   4910: 'Spare_Fault_4910', class No Acknowledgement, trigger "DB302_HMI_Faults_Carrier76_Faults_2" bit 13
   4911: 'Spare_Fault_4911', class No Acknowledgement, trigger "DB302_HMI_Faults_Carrier76_Faults_2" bit 14
   4912: 'Spare_Fault_4912', class No Acknowledgement, trigger "DB302_HMI_Faults_Carrier76_Faults_2" bit 15
   4913: 'Spare_Fault_4913', class No Acknowledgement, trigger "DB302_HMI_Faults_Carrier76_Faults_3" bit 0
   4914: 'Spare_Fault_4914', class No Acknowledgement, trigger "DB302_HMI_Faults_Carrier76_Faults_3" bit 1
   4915: 'Spare_Fault_4915', class No Acknowledgement, trigger "DB302_HMI_Faults_Carrier76_Faults_3" bit 2
   4916: 'Spare_Fault_4916', class No Acknowledgement, trigger "DB302_HMI_Faults_Carrier76_Faults_3" bit 3
   4917: 'Spare_Fault_4917', class No Acknowledgement, trigger "DB302_HMI_Faults_Carrier76_Faults_3" bit 4
   4918: 'Spare_Fault_4918', class No Acknowledgement, trigger "DB302_HMI_Faults_Carrier76_Faults_3" bit 5
   4919: 'Spare_Fault_4919', class No Acknowledgement, trigger "DB302_HMI_Faults_Carrier76_Faults_3" bit 6
   4920: 'Spare_Fault_4920', class No Acknowledgement, trigger "DB302_HMI_Faults_Carrier76_Faults_3" bit 7
   4921: 'Spare_Fault_4921', class No Acknowledgement, trigger "DB302_HMI_Faults_Carrier76_Faults_3" bit 8
   4922: 'Spare_Fault_4922', class No Acknowledgement, trigger "DB302_HMI_Faults_Carrier76_Faults_3" bit 9
   4923: 'Spare_Fault_4923', class No Acknowledgement, trigger "DB302_HMI_Faults_Carrier76_Faults_3" bit 10
   4924: 'Spare_Fault_4924', class No Acknowledgement, trigger "DB302_HMI_Faults_Carrier76_Faults_3" bit 11
   4925: 'Spare_Fault_4925', class No Acknowledgement, trigger "DB302_HMI_Faults_Carrier76_Faults_3" bit 12
   4926: 'Spare_Fault_4926', class No Acknowledgement, trigger "DB302_HMI_Faults_Carrier76_Faults_3" bit 13
   4927: 'Spare_Fault_4927', class No Acknowledgement, trigger "DB302_HMI_Faults_Carrier76_Faults_3" bit 14
   4928: 'Spare_Fault_4928', class No Acknowledgement, trigger "DB302_HMI_Faults_Carrier76_Faults_3" bit 15
   4929: 'Carrier 77 Disconnect Open Power Fault DI11.0', class No Acknowledgement, trigger "DB302_HMI_Faults_Carrier77_Faults_0" bit 0
   4930: 'Carrier 77 Drive Profinet Comm Fault', class No Acknowledgement, trigger "DB302_HMI_Faults_Carrier77_Faults_0" bit 1
   4931: 'Carrier 77 Production Stop Not Reset', class No Acknowledgement, trigger "DB302_HMI_Faults_Carrier77_Faults_0" bit 2
   4932: 'Carrier 77 CB02122 Tripped', class No Acknowledgement, trigger "DB302_HMI_Faults_Carrier77_Faults_0" bit 3
   4933: 'Carrier 77 CB02123 Tripped', class No Acknowledgement, trigger "DB302_HMI_Faults_Carrier77_Faults_0" bit 4
   4934: 'Carrier 77 AUX1 CB Tripped', class No Acknowledgement, trigger "DB302_HMI_Faults_Carrier77_Faults_0" bit 5
   4935: 'Carrier 77 AUX2 CB Tripped', class No Acknowledgement, trigger "DB302_HMI_Faults_Carrier77_Faults_0" bit 6
   4936: 'Carrier 77 PLC Not Communicating', class No Acknowledgement, trigger "DB302_HMI_Faults_Carrier77_Faults_0" bit 7
   4937: 'Carrier 77 Safe Input Card Fault', class No Acknowledgement, trigger "DB302_HMI_Faults_Carrier77_Faults_0" bit 8
   4938: 'Carrier 77 Safe Output Card Fault', class No Acknowledgement, trigger "DB302_HMI_Faults_Carrier77_Faults_0" bit 9
   4939: 'Carrier 77 Standard Input Card Fault', class No Acknowledgement, trigger "DB302_HMI_Faults_Carrier77_Faults_0" bit 10
   4940: 'Carrier 77 Standard Output Card Fault', class No Acknowledgement, trigger "DB302_HMI_Faults_Carrier77_Faults_0" bit 11
   4941: 'Carrier 77 Encoder Position Fault', class No Acknowledgement, trigger "DB302_HMI_Faults_Carrier77_Faults_0" bit 12
   4942: 'Carrier 77 Encoder Internal Error', class No Acknowledgement, trigger "DB302_HMI_Faults_Carrier77_Faults_0" bit 13
   4943: 'Carrier 77 Encoder Comm Fault', class No Acknowledgement, trigger "DB302_HMI_Faults_Carrier77_Faults_0" bit 14
   4944: 'Carrier 77 HMI Comm Fault', class No Acknowledgement, trigger "DB302_HMI_Faults_Carrier77_Faults_0" bit 15
   4945: 'Carrier 77 Crash Detection Fault', class No Acknowledgement, trigger "DB302_HMI_Faults_Carrier77_Faults_1" bit 0
   4946: 'Carrier 77 Carrier Number Invalid', class No Acknowledgement, trigger "DB302_HMI_Faults_Carrier77_Faults_1" bit 1
   4947: 'Carrier 77 Drive: PROFINET configuration error', class No Acknowledgement, trigger "DB302_HMI_Faults_Carrier77_Faults_1" bit 2
   4948: 'Carrier 77 Drive: Error internal communications', class No Acknowledgement, trigger "DB302_HMI_Faults_Carrier77_Faults_1" bit 3
   4949: 'Carrier 77 Drive: Motor overtemperature', class No Acknowledgement, trigger "DB302_HMI_Faults_Carrier77_Faults_1" bit 4
   4950: 'Carrier 77 Drive: Motor overcurrent', class No Acknowledgement, trigger "DB302_HMI_Faults_Carrier77_Faults_1" bit 5
   4951: 'Carrier 77 Drive: Infeed or power unit not ready', class No Acknowledgement, trigger "DB302_HMI_Faults_Carrier77_Faults_1" bit 6
   4952: 'Carrier 77 Drive: Short-circuit/ground fault detected', class No Acknowledgement, trigger "DB302_HMI_Faults_Carrier77_Faults_1" bit 7
   4953: 'Carrier 77 Drive: PROFINET Setpoint timeout', class No Acknowledgement, trigger "DB302_HMI_Faults_Carrier77_Faults_1" bit 8
   4954: 'Carrier 77 Power unit: Overcurrent', class No Acknowledgement, trigger "DB302_HMI_Faults_Carrier77_Faults_1" bit 9
   4955: 'Carrier 77 Power unit: DC link voltage overvoltage', class No Acknowledgement, trigger "DB302_HMI_Faults_Carrier77_Faults_1" bit 10
   4956: 'Carrier 77 Power unit: DC link voltage undervoltage', class No Acknowledgement, trigger "DB302_HMI_Faults_Carrier77_Faults_1" bit 11
   4957: 'Carrier 77 Power unit: Line phase failure in main circuit', class No Acknowledgement, trigger "DB302_HMI_Faults_Carrier77_Faults_1" bit 12
   4958: 'Carrier 77 Power unit: Phase failure motor cable', class No Acknowledgement, trigger "DB302_HMI_Faults_Carrier77_Faults_1" bit 13
   4959: 'Carrier 77 Power unit: Ground fault', class No Acknowledgement, trigger "DB302_HMI_Faults_Carrier77_Faults_1" bit 14
   4960: 'Spare_Fault_4960', class No Acknowledgement, trigger "DB302_HMI_Faults_Carrier77_Faults_1" bit 15
   4961: 'Carrier 77 Motion Off Fault', class No Acknowledgement, trigger "DB302_HMI_Faults_Carrier77_Faults_2" bit 0
   4962: 'Carrier 77 Motion On Fault', class No Acknowledgement, trigger "DB302_HMI_Faults_Carrier77_Faults_2" bit 1
   4963: 'Carrier 77 Spacing Fault', class No Acknowledgement, trigger "DB302_HMI_Faults_Carrier77_Faults_2" bit 2
   4964: 'Carrier 77 Duplicate Carrier Number Fault', class No Acknowledgement, trigger "DB302_HMI_Faults_Carrier77_Faults_2" bit 3
   4965: 'Spare_Fault_4965', class No Acknowledgement, trigger "DB302_HMI_Faults_Carrier77_Faults_2" bit 4
   4966: 'Spare_Fault_4966', class No Acknowledgement, trigger "DB302_HMI_Faults_Carrier77_Faults_2" bit 5
   4967: 'Spare_Fault_4967', class No Acknowledgement, trigger "DB302_HMI_Faults_Carrier77_Faults_2" bit 6
   4968: 'Spare_Fault_4968', class No Acknowledgement, trigger "DB302_HMI_Faults_Carrier77_Faults_2" bit 7
   4969: 'Spare_Fault_4969', class No Acknowledgement, trigger "DB302_HMI_Faults_Carrier77_Faults_2" bit 8
   4970: 'Spare_Fault_4970', class No Acknowledgement, trigger "DB302_HMI_Faults_Carrier77_Faults_2" bit 9
   4971: 'Spare_Fault_4971', class No Acknowledgement, trigger "DB302_HMI_Faults_Carrier77_Faults_2" bit 10
   4972: 'Spare_Fault_4972', class No Acknowledgement, trigger "DB302_HMI_Faults_Carrier77_Faults_2" bit 11
   4973: 'Spare_Fault_4973', class No Acknowledgement, trigger "DB302_HMI_Faults_Carrier77_Faults_2" bit 12
   4974: 'Spare_Fault_4974', class No Acknowledgement, trigger "DB302_HMI_Faults_Carrier77_Faults_2" bit 13
   4975: 'Spare_Fault_4975', class No Acknowledgement, trigger "DB302_HMI_Faults_Carrier77_Faults_2" bit 14
   4976: 'Spare_Fault_4976', class No Acknowledgement, trigger "DB302_HMI_Faults_Carrier77_Faults_2" bit 15
   4977: 'Spare_Fault_4977', class No Acknowledgement, trigger "DB302_HMI_Faults_Carrier77_Faults_3" bit 0
   4978: 'Spare_Fault_4978', class No Acknowledgement, trigger "DB302_HMI_Faults_Carrier77_Faults_3" bit 1
   4979: 'Spare_Fault_4979', class No Acknowledgement, trigger "DB302_HMI_Faults_Carrier77_Faults_3" bit 2
   4980: 'Spare_Fault_4980', class No Acknowledgement, trigger "DB302_HMI_Faults_Carrier77_Faults_3" bit 3
   4981: 'Spare_Fault_4981', class No Acknowledgement, trigger "DB302_HMI_Faults_Carrier77_Faults_3" bit 4
   4982: 'Spare_Fault_4982', class No Acknowledgement, trigger "DB302_HMI_Faults_Carrier77_Faults_3" bit 5
   4983: 'Spare_Fault_4983', class No Acknowledgement, trigger "DB302_HMI_Faults_Carrier77_Faults_3" bit 6
   4984: 'Spare_Fault_4984', class No Acknowledgement, trigger "DB302_HMI_Faults_Carrier77_Faults_3" bit 7
   4985: 'Spare_Fault_4985', class No Acknowledgement, trigger "DB302_HMI_Faults_Carrier77_Faults_3" bit 8
   4986: 'Spare_Fault_4986', class No Acknowledgement, trigger "DB302_HMI_Faults_Carrier77_Faults_3" bit 9
   4987: 'Spare_Fault_4987', class No Acknowledgement, trigger "DB302_HMI_Faults_Carrier77_Faults_3" bit 10
   4988: 'Spare_Fault_4988', class No Acknowledgement, trigger "DB302_HMI_Faults_Carrier77_Faults_3" bit 11
   4989: 'Spare_Fault_4989', class No Acknowledgement, trigger "DB302_HMI_Faults_Carrier77_Faults_3" bit 12
   4990: 'Spare_Fault_4990', class No Acknowledgement, trigger "DB302_HMI_Faults_Carrier77_Faults_3" bit 13
   4991: 'Spare_Fault_4991', class No Acknowledgement, trigger "DB302_HMI_Faults_Carrier77_Faults_3" bit 14
   4992: 'Spare_Fault_4992', class No Acknowledgement, trigger "DB302_HMI_Faults_Carrier77_Faults_3" bit 15
   4993: 'Carrier 78 Disconnect Open Power Fault DI11.0', class No Acknowledgement, trigger "DB302_HMI_Faults_Carrier78_Faults_0" bit 0
   4994: 'Carrier 78 Drive Profinet Comm Fault', class No Acknowledgement, trigger "DB302_HMI_Faults_Carrier78_Faults_0" bit 1
   4995: 'Carrier 78 Production Stop Not Reset', class No Acknowledgement, trigger "DB302_HMI_Faults_Carrier78_Faults_0" bit 2
   4996: 'Carrier 78 CB02122 Tripped', class No Acknowledgement, trigger "DB302_HMI_Faults_Carrier78_Faults_0" bit 3
   4997: 'Carrier 78 CB02123 Tripped', class No Acknowledgement, trigger "DB302_HMI_Faults_Carrier78_Faults_0" bit 4
   4998: 'Carrier 78 AUX1 CB Tripped', class No Acknowledgement, trigger "DB302_HMI_Faults_Carrier78_Faults_0" bit 5
   4999: 'Carrier 78 AUX2 CB Tripped', class No Acknowledgement, trigger "DB302_HMI_Faults_Carrier78_Faults_0" bit 6
   5000: 'Carrier 78 PLC Not Communicating', class No Acknowledgement, trigger "DB302_HMI_Faults_Carrier78_Faults_0" bit 7
   5001: 'Carrier 78 Safe Input Card Fault', class No Acknowledgement, trigger "DB302_HMI_Faults_Carrier78_Faults_0" bit 8
   5002: 'Carrier 78 Safe Output Card Fault', class No Acknowledgement, trigger "DB302_HMI_Faults_Carrier78_Faults_0" bit 9
   5003: 'Carrier 78 Standard Input Card Fault', class No Acknowledgement, trigger "DB302_HMI_Faults_Carrier78_Faults_0" bit 10
   5004: 'Carrier 78 Standard Output Card Fault', class No Acknowledgement, trigger "DB302_HMI_Faults_Carrier78_Faults_0" bit 11
   5005: 'Carrier 78 Encoder Position Fault', class No Acknowledgement, trigger "DB302_HMI_Faults_Carrier78_Faults_0" bit 12
   5006: 'Carrier 78 Encoder Internal Error', class No Acknowledgement, trigger "DB302_HMI_Faults_Carrier78_Faults_0" bit 13
   5007: 'Carrier 78 Encoder Comm Fault', class No Acknowledgement, trigger "DB302_HMI_Faults_Carrier78_Faults_0" bit 14
   5008: 'Carrier 78 HMI Comm Fault', class No Acknowledgement, trigger "DB302_HMI_Faults_Carrier78_Faults_0" bit 15
   5009: 'Carrier 78 Crash Detection Fault', class No Acknowledgement, trigger "DB302_HMI_Faults_Carrier78_Faults_1" bit 0
   5010: 'Carrier 78 Carrier Number Invalid', class No Acknowledgement, trigger "DB302_HMI_Faults_Carrier78_Faults_1" bit 1
   5011: 'Carrier 78 Drive: PROFINET configuration error', class No Acknowledgement, trigger "DB302_HMI_Faults_Carrier78_Faults_1" bit 2
   5012: 'Carrier 78 Drive: Error internal communications', class No Acknowledgement, trigger "DB302_HMI_Faults_Carrier78_Faults_1" bit 3
   5013: 'Carrier 78 Drive: Motor overtemperature', class No Acknowledgement, trigger "DB302_HMI_Faults_Carrier78_Faults_1" bit 4
   5014: 'Carrier 78 Drive: Motor overcurrent', class No Acknowledgement, trigger "DB302_HMI_Faults_Carrier78_Faults_1" bit 5
   5015: 'Carrier 78 Drive: Infeed or power unit not ready', class No Acknowledgement, trigger "DB302_HMI_Faults_Carrier78_Faults_1" bit 6
   5016: 'Carrier 78 Drive: Short-circuit/ground fault detected', class No Acknowledgement, trigger "DB302_HMI_Faults_Carrier78_Faults_1" bit 7
   5017: 'Carrier 78 Drive: PROFINET Setpoint timeout', class No Acknowledgement, trigger "DB302_HMI_Faults_Carrier78_Faults_1" bit 8
   5018: 'Carrier 78 Power unit: Overcurrent', class No Acknowledgement, trigger "DB302_HMI_Faults_Carrier78_Faults_1" bit 9
   5019: 'Carrier 78 Power unit: DC link voltage overvoltage', class No Acknowledgement, trigger "DB302_HMI_Faults_Carrier78_Faults_1" bit 10
   5020: 'Carrier 78 Power unit: DC link voltage undervoltage', class No Acknowledgement, trigger "DB302_HMI_Faults_Carrier78_Faults_1" bit 11
   5021: 'Carrier 78 Power unit: Line phase failure in main circuit', class No Acknowledgement, trigger "DB302_HMI_Faults_Carrier78_Faults_1" bit 12
   5022: 'Carrier 78 Power unit: Phase failure motor cable', class No Acknowledgement, trigger "DB302_HMI_Faults_Carrier78_Faults_1" bit 13
   5023: 'Carrier 78 Power unit: Ground fault', class No Acknowledgement, trigger "DB302_HMI_Faults_Carrier78_Faults_1" bit 14
   5024: 'Spare_Fault_5024', class No Acknowledgement, trigger "DB302_HMI_Faults_Carrier78_Faults_1" bit 15
   5025: 'Carrier 78 Motion Off Fault', class No Acknowledgement, trigger "DB302_HMI_Faults_Carrier78_Faults_2" bit 0
   5026: 'Carrier 78 Motion On Fault', class No Acknowledgement, trigger "DB302_HMI_Faults_Carrier78_Faults_2" bit 1
   5027: 'Carrier 78 Spacing Fault', class No Acknowledgement, trigger "DB302_HMI_Faults_Carrier78_Faults_2" bit 2
   5028: 'Carrier 78 Duplicate Carrier Number Fault', class No Acknowledgement, trigger "DB302_HMI_Faults_Carrier78_Faults_2" bit 3
   5029: 'Spare_Fault_5029', class No Acknowledgement, trigger "DB302_HMI_Faults_Carrier78_Faults_2" bit 4
   5030: 'Spare_Fault_5030', class No Acknowledgement, trigger "DB302_HMI_Faults_Carrier78_Faults_2" bit 5
   5031: 'Spare_Fault_5031', class No Acknowledgement, trigger "DB302_HMI_Faults_Carrier78_Faults_2" bit 6
   5032: 'Spare_Fault_5032', class No Acknowledgement, trigger "DB302_HMI_Faults_Carrier78_Faults_2" bit 7
   5033: 'Spare_Fault_5033', class No Acknowledgement, trigger "DB302_HMI_Faults_Carrier78_Faults_2" bit 8
   5034: 'Spare_Fault_5034', class No Acknowledgement, trigger "DB302_HMI_Faults_Carrier78_Faults_2" bit 9
   5035: 'Spare_Fault_5035', class No Acknowledgement, trigger "DB302_HMI_Faults_Carrier78_Faults_2" bit 10
   5036: 'Spare_Fault_5036', class No Acknowledgement, trigger "DB302_HMI_Faults_Carrier78_Faults_2" bit 11
   5037: 'Spare_Fault_5037', class No Acknowledgement, trigger "DB302_HMI_Faults_Carrier78_Faults_2" bit 12
   5038: 'Spare_Fault_5038', class No Acknowledgement, trigger "DB302_HMI_Faults_Carrier78_Faults_2" bit 13
   5039: 'Spare_Fault_5039', class No Acknowledgement, trigger "DB302_HMI_Faults_Carrier78_Faults_2" bit 14
   5040: 'Spare_Fault_5040', class No Acknowledgement, trigger "DB302_HMI_Faults_Carrier78_Faults_2" bit 15
   5041: 'Spare_Fault_5041', class No Acknowledgement, trigger "DB302_HMI_Faults_Carrier78_Faults_3" bit 0
   5042: 'Spare_Fault_5042', class No Acknowledgement, trigger "DB302_HMI_Faults_Carrier78_Faults_3" bit 1
   5043: 'Spare_Fault_5043', class No Acknowledgement, trigger "DB302_HMI_Faults_Carrier78_Faults_3" bit 2
   5044: 'Spare_Fault_5044', class No Acknowledgement, trigger "DB302_HMI_Faults_Carrier78_Faults_3" bit 3
   5045: 'Spare_Fault_5045', class No Acknowledgement, trigger "DB302_HMI_Faults_Carrier78_Faults_3" bit 4
   5046: 'Spare_Fault_5046', class No Acknowledgement, trigger "DB302_HMI_Faults_Carrier78_Faults_3" bit 5
   5047: 'Spare_Fault_5047', class No Acknowledgement, trigger "DB302_HMI_Faults_Carrier78_Faults_3" bit 6
   5048: 'Spare_Fault_5048', class No Acknowledgement, trigger "DB302_HMI_Faults_Carrier78_Faults_3" bit 7
   5049: 'Spare_Fault_5049', class No Acknowledgement, trigger "DB302_HMI_Faults_Carrier78_Faults_3" bit 8
   5050: 'Spare_Fault_5050', class No Acknowledgement, trigger "DB302_HMI_Faults_Carrier78_Faults_3" bit 9
   5051: 'Spare_Fault_5051', class No Acknowledgement, trigger "DB302_HMI_Faults_Carrier78_Faults_3" bit 10
   5052: 'Spare_Fault_5052', class No Acknowledgement, trigger "DB302_HMI_Faults_Carrier78_Faults_3" bit 11
   5053: 'Spare_Fault_5053', class No Acknowledgement, trigger "DB302_HMI_Faults_Carrier78_Faults_3" bit 12
   5054: 'Spare_Fault_5054', class No Acknowledgement, trigger "DB302_HMI_Faults_Carrier78_Faults_3" bit 13
   5055: 'Spare_Fault_5055', class No Acknowledgement, trigger "DB302_HMI_Faults_Carrier78_Faults_3" bit 14
   5056: 'Spare_Fault_5056', class No Acknowledgement, trigger "DB302_HMI_Faults_Carrier78_Faults_3" bit 15
   5057: 'Carrier 79 Disconnect Open Power Fault DI11.0', class No Acknowledgement, trigger "DB302_HMI_Faults_Carrier79_Faults_0" bit 0
   5058: 'Carrier 79 Drive Profinet Comm Fault', class No Acknowledgement, trigger "DB302_HMI_Faults_Carrier79_Faults_0" bit 1
   5059: 'Carrier 79 Production Stop Not Reset', class No Acknowledgement, trigger "DB302_HMI_Faults_Carrier79_Faults_0" bit 2
   5060: 'Carrier 79 CB02122 Tripped', class No Acknowledgement, trigger "DB302_HMI_Faults_Carrier79_Faults_0" bit 3
   5061: 'Carrier 79 CB02123 Tripped', class No Acknowledgement, trigger "DB302_HMI_Faults_Carrier79_Faults_0" bit 4
   5062: 'Carrier 79 AUX1 CB Tripped', class No Acknowledgement, trigger "DB302_HMI_Faults_Carrier79_Faults_0" bit 5
   5063: 'Carrier 79 AUX2 CB Tripped', class No Acknowledgement, trigger "DB302_HMI_Faults_Carrier79_Faults_0" bit 6
   5064: 'Carrier 79 PLC Not Communicating', class No Acknowledgement, trigger "DB302_HMI_Faults_Carrier79_Faults_0" bit 7
   5065: 'Carrier 79 Safe Input Card Fault', class No Acknowledgement, trigger "DB302_HMI_Faults_Carrier79_Faults_0" bit 8
   5066: 'Carrier 79 Safe Output Card Fault', class No Acknowledgement, trigger "DB302_HMI_Faults_Carrier79_Faults_0" bit 9
   5067: 'Carrier 79 Standard Input Card Fault', class No Acknowledgement, trigger "DB302_HMI_Faults_Carrier79_Faults_0" bit 10
   5068: 'Carrier 79 Standard Output Card Fault', class No Acknowledgement, trigger "DB302_HMI_Faults_Carrier79_Faults_0" bit 11
   5069: 'Carrier 79 Encoder Position Fault', class No Acknowledgement, trigger "DB302_HMI_Faults_Carrier79_Faults_0" bit 12
   5070: 'Carrier 79 Encoder Internal Error', class No Acknowledgement, trigger "DB302_HMI_Faults_Carrier79_Faults_0" bit 13
   5071: 'Carrier 79 Encoder Comm Fault', class No Acknowledgement, trigger "DB302_HMI_Faults_Carrier79_Faults_0" bit 14
   5072: 'Carrier 79 HMI Comm Fault', class No Acknowledgement, trigger "DB302_HMI_Faults_Carrier79_Faults_0" bit 15
   5073: 'Carrier 79 Crash Detection Fault', class No Acknowledgement, trigger "DB302_HMI_Faults_Carrier79_Faults_1" bit 0
   5074: 'Carrier 79 Carrier Number Invalid', class No Acknowledgement, trigger "DB302_HMI_Faults_Carrier79_Faults_1" bit 1
   5075: 'Carrier 79 Drive: PROFINET configuration error', class No Acknowledgement, trigger "DB302_HMI_Faults_Carrier79_Faults_1" bit 2
   5076: 'Carrier 79 Drive: Error internal communications', class No Acknowledgement, trigger "DB302_HMI_Faults_Carrier79_Faults_1" bit 3
   5077: 'Carrier 79 Drive: Motor overtemperature', class No Acknowledgement, trigger "DB302_HMI_Faults_Carrier79_Faults_1" bit 4
   5078: 'Carrier 79 Drive: Motor overcurrent', class No Acknowledgement, trigger "DB302_HMI_Faults_Carrier79_Faults_1" bit 5
   5079: 'Carrier 79 Drive: Infeed or power unit not ready', class No Acknowledgement, trigger "DB302_HMI_Faults_Carrier79_Faults_1" bit 6
   5080: 'Carrier 79 Drive: Short-circuit/ground fault detected', class No Acknowledgement, trigger "DB302_HMI_Faults_Carrier79_Faults_1" bit 7
   5081: 'Carrier 79 Drive: PROFINET Setpoint timeout', class No Acknowledgement, trigger "DB302_HMI_Faults_Carrier79_Faults_1" bit 8
   5082: 'Carrier 79 Power unit: Overcurrent', class No Acknowledgement, trigger "DB302_HMI_Faults_Carrier79_Faults_1" bit 9
   5083: 'Carrier 79 Power unit: DC link voltage overvoltage', class No Acknowledgement, trigger "DB302_HMI_Faults_Carrier79_Faults_1" bit 10
   5084: 'Carrier 79 Power unit: DC link voltage undervoltage', class No Acknowledgement, trigger "DB302_HMI_Faults_Carrier79_Faults_1" bit 11
   5085: 'Carrier 79 Power unit: Line phase failure in main circuit', class No Acknowledgement, trigger "DB302_HMI_Faults_Carrier79_Faults_1" bit 12
   5086: 'Carrier 79 Power unit: Phase failure motor cable', class No Acknowledgement, trigger "DB302_HMI_Faults_Carrier79_Faults_1" bit 13
   5087: 'Carrier 79 Power unit: Ground fault', class No Acknowledgement, trigger "DB302_HMI_Faults_Carrier79_Faults_1" bit 14
   5088: 'Spare_Fault_5088', class No Acknowledgement, trigger "DB302_HMI_Faults_Carrier79_Faults_1" bit 15
   5089: 'Carrier 79 Motion Off Fault', class No Acknowledgement, trigger "DB302_HMI_Faults_Carrier79_Faults_2" bit 0
   5090: 'Carrier 79 Motion On Fault', class No Acknowledgement, trigger "DB302_HMI_Faults_Carrier79_Faults_2" bit 1
   5091: 'Carrier 79 Spacing Fault', class No Acknowledgement, trigger "DB302_HMI_Faults_Carrier79_Faults_2" bit 2
   5092: 'Carrier 79 Duplicate Carrier Number Fault', class No Acknowledgement, trigger "DB302_HMI_Faults_Carrier79_Faults_2" bit 3
   5093: 'Spare_Fault_5093', class No Acknowledgement, trigger "DB302_HMI_Faults_Carrier79_Faults_2" bit 4
   5094: 'Spare_Fault_5094', class No Acknowledgement, trigger "DB302_HMI_Faults_Carrier79_Faults_2" bit 5
   5095: 'Spare_Fault_5095', class No Acknowledgement, trigger "DB302_HMI_Faults_Carrier79_Faults_2" bit 6
   5096: 'Spare_Fault_5096', class No Acknowledgement, trigger "DB302_HMI_Faults_Carrier79_Faults_2" bit 7
   5097: 'Spare_Fault_5097', class No Acknowledgement, trigger "DB302_HMI_Faults_Carrier79_Faults_2" bit 8
   5098: 'Spare_Fault_5098', class No Acknowledgement, trigger "DB302_HMI_Faults_Carrier79_Faults_2" bit 9
   5099: 'Spare_Fault_5099', class No Acknowledgement, trigger "DB302_HMI_Faults_Carrier79_Faults_2" bit 10
   5100: 'Spare_Fault_5100', class No Acknowledgement, trigger "DB302_HMI_Faults_Carrier79_Faults_2" bit 11
   5101: 'Spare_Fault_5101', class No Acknowledgement, trigger "DB302_HMI_Faults_Carrier79_Faults_2" bit 12
   5102: 'Spare_Fault_5102', class No Acknowledgement, trigger "DB302_HMI_Faults_Carrier79_Faults_2" bit 13
   5103: 'Spare_Fault_5103', class No Acknowledgement, trigger "DB302_HMI_Faults_Carrier79_Faults_2" bit 14
   5104: 'Spare_Fault_5104', class No Acknowledgement, trigger "DB302_HMI_Faults_Carrier79_Faults_2" bit 15
   5105: 'Spare_Fault_5105', class No Acknowledgement, trigger "DB302_HMI_Faults_Carrier79_Faults_3" bit 0
   5106: 'Spare_Fault_5106', class No Acknowledgement, trigger "DB302_HMI_Faults_Carrier79_Faults_3" bit 1
   5107: 'Spare_Fault_5107', class No Acknowledgement, trigger "DB302_HMI_Faults_Carrier79_Faults_3" bit 2
   5108: 'Spare_Fault_5108', class No Acknowledgement, trigger "DB302_HMI_Faults_Carrier79_Faults_3" bit 3
   5109: 'Spare_Fault_5109', class No Acknowledgement, trigger "DB302_HMI_Faults_Carrier79_Faults_3" bit 4
   5110: 'Spare_Fault_5110', class No Acknowledgement, trigger "DB302_HMI_Faults_Carrier79_Faults_3" bit 5
   5111: 'Spare_Fault_5111', class No Acknowledgement, trigger "DB302_HMI_Faults_Carrier79_Faults_3" bit 6
   5112: 'Spare_Fault_5112', class No Acknowledgement, trigger "DB302_HMI_Faults_Carrier79_Faults_3" bit 7
   5113: 'Spare_Fault_5113', class No Acknowledgement, trigger "DB302_HMI_Faults_Carrier79_Faults_3" bit 8
   5114: 'Spare_Fault_5114', class No Acknowledgement, trigger "DB302_HMI_Faults_Carrier79_Faults_3" bit 9
   5115: 'Spare_Fault_5115', class No Acknowledgement, trigger "DB302_HMI_Faults_Carrier79_Faults_3" bit 10
   5116: 'Spare_Fault_5116', class No Acknowledgement, trigger "DB302_HMI_Faults_Carrier79_Faults_3" bit 11
   5117: 'Spare_Fault_5117', class No Acknowledgement, trigger "DB302_HMI_Faults_Carrier79_Faults_3" bit 12
   5118: 'Spare_Fault_5118', class No Acknowledgement, trigger "DB302_HMI_Faults_Carrier79_Faults_3" bit 13
   5119: 'Spare_Fault_5119', class No Acknowledgement, trigger "DB302_HMI_Faults_Carrier79_Faults_3" bit 14
   5120: 'Spare_Fault_5120', class No Acknowledgement, trigger "DB302_HMI_Faults_Carrier79_Faults_3" bit 15
   5121: 'Carrier 80 Disconnect Open Power Fault DI11.0', class No Acknowledgement, trigger "DB302_HMI_Faults_Carrier80_Faults_0" bit 0
   5122: 'Carrier 80 Drive Profinet Comm Fault', class No Acknowledgement, trigger "DB302_HMI_Faults_Carrier80_Faults_0" bit 1
   5123: 'Carrier 80 Production Stop Not Reset', class No Acknowledgement, trigger "DB302_HMI_Faults_Carrier80_Faults_0" bit 2
   5124: 'Carrier 80 CB02122 Tripped', class No Acknowledgement, trigger "DB302_HMI_Faults_Carrier80_Faults_0" bit 3
   5125: 'Carrier 80 CB02123 Tripped', class No Acknowledgement, trigger "DB302_HMI_Faults_Carrier80_Faults_0" bit 4
   5126: 'Carrier 80 AUX1 CB Tripped', class No Acknowledgement, trigger "DB302_HMI_Faults_Carrier80_Faults_0" bit 5
   5127: 'Carrier 80 AUX2 CB Tripped', class No Acknowledgement, trigger "DB302_HMI_Faults_Carrier80_Faults_0" bit 6
   5128: 'Carrier 80 PLC Not Communicating', class No Acknowledgement, trigger "DB302_HMI_Faults_Carrier80_Faults_0" bit 7
   5129: 'Carrier 80 Safe Input Card Fault', class No Acknowledgement, trigger "DB302_HMI_Faults_Carrier80_Faults_0" bit 8
   5130: 'Carrier 80 Safe Output Card Fault', class No Acknowledgement, trigger "DB302_HMI_Faults_Carrier80_Faults_0" bit 9
   5131: 'Carrier 80 Standard Input Card Fault', class No Acknowledgement, trigger "DB302_HMI_Faults_Carrier80_Faults_0" bit 10
   5132: 'Carrier 80 Standard Output Card Fault', class No Acknowledgement, trigger "DB302_HMI_Faults_Carrier80_Faults_0" bit 11
   5133: 'Carrier 80 Encoder Position Fault', class No Acknowledgement, trigger "DB302_HMI_Faults_Carrier80_Faults_0" bit 12
   5134: 'Carrier 80 Encoder Internal Error', class No Acknowledgement, trigger "DB302_HMI_Faults_Carrier80_Faults_0" bit 13
   5135: 'Carrier 80 Encoder Comm Fault', class No Acknowledgement, trigger "DB302_HMI_Faults_Carrier80_Faults_0" bit 14
   5136: 'Carrier 80 HMI Comm Fault', class No Acknowledgement, trigger "DB302_HMI_Faults_Carrier80_Faults_0" bit 15
   5137: 'Carrier 80 Crash Detection Fault', class No Acknowledgement, trigger "DB302_HMI_Faults_Carrier80_Faults_1" bit 0
   5138: 'Carrier 80 Carrier Number Invalid', class No Acknowledgement, trigger "DB302_HMI_Faults_Carrier80_Faults_1" bit 1
   5139: 'Carrier 80 Drive: PROFINET configuration error', class No Acknowledgement, trigger "DB302_HMI_Faults_Carrier80_Faults_1" bit 2
   5140: 'Carrier 80 Drive: Error internal communications', class No Acknowledgement, trigger "DB302_HMI_Faults_Carrier80_Faults_1" bit 3
   5141: 'Carrier 80 Drive: Motor overtemperature', class No Acknowledgement, trigger "DB302_HMI_Faults_Carrier80_Faults_1" bit 4
   5142: 'Carrier 80 Drive: Motor overcurrent', class No Acknowledgement, trigger "DB302_HMI_Faults_Carrier80_Faults_1" bit 5
   5143: 'Carrier 80 Drive: Infeed or power unit not ready', class No Acknowledgement, trigger "DB302_HMI_Faults_Carrier80_Faults_1" bit 6
   5144: 'Carrier 80 Drive: Short-circuit/ground fault detected', class No Acknowledgement, trigger "DB302_HMI_Faults_Carrier80_Faults_1" bit 7
   5145: 'Carrier 80 Drive: PROFINET Setpoint timeout', class No Acknowledgement, trigger "DB302_HMI_Faults_Carrier80_Faults_1" bit 8
   5146: 'Carrier 80 Power unit: Overcurrent', class No Acknowledgement, trigger "DB302_HMI_Faults_Carrier80_Faults_1" bit 9
   5147: 'Carrier 80 Power unit: DC link voltage overvoltage', class No Acknowledgement, trigger "DB302_HMI_Faults_Carrier80_Faults_1" bit 10
   5148: 'Carrier 80 Power unit: DC link voltage undervoltage', class No Acknowledgement, trigger "DB302_HMI_Faults_Carrier80_Faults_1" bit 11
   5149: 'Carrier 80 Power unit: Line phase failure in main circuit', class No Acknowledgement, trigger "DB302_HMI_Faults_Carrier80_Faults_1" bit 12
   5150: 'Carrier 80 Power unit: Phase failure motor cable', class No Acknowledgement, trigger "DB302_HMI_Faults_Carrier80_Faults_1" bit 13
   5151: 'Carrier 80 Power unit: Ground fault', class No Acknowledgement, trigger "DB302_HMI_Faults_Carrier80_Faults_1" bit 14
   5152: 'Spare_Fault_5152', class No Acknowledgement, trigger "DB302_HMI_Faults_Carrier80_Faults_1" bit 15
   5153: 'Carrier 80 Motion Off Fault', class No Acknowledgement, trigger "DB302_HMI_Faults_Carrier80_Faults_2" bit 0
   5154: 'Carrier 80 Motion On Fault', class No Acknowledgement, trigger "DB302_HMI_Faults_Carrier80_Faults_2" bit 1
   5155: 'Carrier 80 Spacing Fault', class No Acknowledgement, trigger "DB302_HMI_Faults_Carrier80_Faults_2" bit 2
   5156: 'Carrier 80 Duplicate Carrier Number Fault', class No Acknowledgement, trigger "DB302_HMI_Faults_Carrier80_Faults_2" bit 3
   5157: 'Spare_Fault_5157', class No Acknowledgement, trigger "DB302_HMI_Faults_Carrier80_Faults_2" bit 4
   5158: 'Spare_Fault_5158', class No Acknowledgement, trigger "DB302_HMI_Faults_Carrier80_Faults_2" bit 5
   5159: 'Spare_Fault_5159', class No Acknowledgement, trigger "DB302_HMI_Faults_Carrier80_Faults_2" bit 6
   5160: 'Spare_Fault_5160', class No Acknowledgement, trigger "DB302_HMI_Faults_Carrier80_Faults_2" bit 7
   5161: 'Spare_Fault_5161', class No Acknowledgement, trigger "DB302_HMI_Faults_Carrier80_Faults_2" bit 8
   5162: 'Spare_Fault_5162', class No Acknowledgement, trigger "DB302_HMI_Faults_Carrier80_Faults_2" bit 9
   5163: 'Spare_Fault_5163', class No Acknowledgement, trigger "DB302_HMI_Faults_Carrier80_Faults_2" bit 10
   5164: 'Spare_Fault_5164', class No Acknowledgement, trigger "DB302_HMI_Faults_Carrier80_Faults_2" bit 11
   5165: 'Spare_Fault_5165', class No Acknowledgement, trigger "DB302_HMI_Faults_Carrier80_Faults_2" bit 12
   5166: 'Spare_Fault_5166', class No Acknowledgement, trigger "DB302_HMI_Faults_Carrier80_Faults_2" bit 13
   5167: 'Spare_Fault_5167', class No Acknowledgement, trigger "DB302_HMI_Faults_Carrier80_Faults_2" bit 14
   5168: 'Spare_Fault_5168', class No Acknowledgement, trigger "DB302_HMI_Faults_Carrier80_Faults_2" bit 15
   5169: 'Spare_Fault_5169', class No Acknowledgement, trigger "DB302_HMI_Faults_Carrier80_Faults_3" bit 0
   5170: 'Spare_Fault_5170', class No Acknowledgement, trigger "DB302_HMI_Faults_Carrier80_Faults_3" bit 1
   5171: 'Spare_Fault_5171', class No Acknowledgement, trigger "DB302_HMI_Faults_Carrier80_Faults_3" bit 2
   5172: 'Spare_Fault_5172', class No Acknowledgement, trigger "DB302_HMI_Faults_Carrier80_Faults_3" bit 3
   5173: 'Spare_Fault_5173', class No Acknowledgement, trigger "DB302_HMI_Faults_Carrier80_Faults_3" bit 4
   5174: 'Spare_Fault_5174', class No Acknowledgement, trigger "DB302_HMI_Faults_Carrier80_Faults_3" bit 5
   5175: 'Spare_Fault_5175', class No Acknowledgement, trigger "DB302_HMI_Faults_Carrier80_Faults_3" bit 6
   5176: 'Spare_Fault_5176', class No Acknowledgement, trigger "DB302_HMI_Faults_Carrier80_Faults_3" bit 7
   5177: 'Spare_Fault_5177', class No Acknowledgement, trigger "DB302_HMI_Faults_Carrier80_Faults_3" bit 8
   5178: 'Spare_Fault_5178', class No Acknowledgement, trigger "DB302_HMI_Faults_Carrier80_Faults_3" bit 9
   5179: 'Spare_Fault_5179', class No Acknowledgement, trigger "DB302_HMI_Faults_Carrier80_Faults_3" bit 10
   5180: 'Spare_Fault_5180', class No Acknowledgement, trigger "DB302_HMI_Faults_Carrier80_Faults_3" bit 11
   5181: 'Spare_Fault_5181', class No Acknowledgement, trigger "DB302_HMI_Faults_Carrier80_Faults_3" bit 12
   5182: 'Spare_Fault_5182', class No Acknowledgement, trigger "DB302_HMI_Faults_Carrier80_Faults_3" bit 13
   5183: 'Spare_Fault_5183', class No Acknowledgement, trigger "DB302_HMI_Faults_Carrier80_Faults_3" bit 14
   5184: 'Spare_Fault_5184', class No Acknowledgement, trigger "DB302_HMI_Faults_Carrier80_Faults_3" bit 15
   5185: 'Carrier 81 Disconnect Open Power Fault DI11.0', class No Acknowledgement, trigger "DB302_HMI_Faults_Carrier81_Faults_0" bit 0
   5186: 'Carrier 81 Drive Profinet Comm Fault', class No Acknowledgement, trigger "DB302_HMI_Faults_Carrier81_Faults_0" bit 1
   5187: 'Carrier 81 Production Stop Not Reset', class No Acknowledgement, trigger "DB302_HMI_Faults_Carrier81_Faults_0" bit 2
   5188: 'Carrier 81 CB02122 Tripped', class No Acknowledgement, trigger "DB302_HMI_Faults_Carrier81_Faults_0" bit 3
   5189: 'Carrier 81 CB02123 Tripped', class No Acknowledgement, trigger "DB302_HMI_Faults_Carrier81_Faults_0" bit 4
   5190: 'Carrier 81 AUX1 CB Tripped', class No Acknowledgement, trigger "DB302_HMI_Faults_Carrier81_Faults_0" bit 5
   5191: 'Carrier 81 AUX2 CB Tripped', class No Acknowledgement, trigger "DB302_HMI_Faults_Carrier81_Faults_0" bit 6
   5192: 'Carrier 81 PLC Not Communicating', class No Acknowledgement, trigger "DB302_HMI_Faults_Carrier81_Faults_0" bit 7
   5193: 'Carrier 81 Safe Input Card Fault', class No Acknowledgement, trigger "DB302_HMI_Faults_Carrier81_Faults_0" bit 8
   5194: 'Carrier 81 Safe Output Card Fault', class No Acknowledgement, trigger "DB302_HMI_Faults_Carrier81_Faults_0" bit 9
   5195: 'Carrier 81 Standard Input Card Fault', class No Acknowledgement, trigger "DB302_HMI_Faults_Carrier81_Faults_0" bit 10
   5196: 'Carrier 81 Standard Output Card Fault', class No Acknowledgement, trigger "DB302_HMI_Faults_Carrier81_Faults_0" bit 11
   5197: 'Carrier 81 Encoder Position Fault', class No Acknowledgement, trigger "DB302_HMI_Faults_Carrier81_Faults_0" bit 12
   5198: 'Carrier 81 Encoder Internal Error', class No Acknowledgement, trigger "DB302_HMI_Faults_Carrier81_Faults_0" bit 13
   5199: 'Carrier 81 Encoder Comm Fault', class No Acknowledgement, trigger "DB302_HMI_Faults_Carrier81_Faults_0" bit 14
   5200: 'Carrier 81 HMI Comm Fault', class No Acknowledgement, trigger "DB302_HMI_Faults_Carrier81_Faults_0" bit 15
   5201: 'Carrier 81 Crash Detection Fault', class No Acknowledgement, trigger "DB302_HMI_Faults_Carrier81_Faults_1" bit 0
   5202: 'Carrier 81 Carrier Number Invalid', class No Acknowledgement, trigger "DB302_HMI_Faults_Carrier81_Faults_1" bit 1
   5203: 'Carrier 81 Drive: PROFINET configuration error', class No Acknowledgement, trigger "DB302_HMI_Faults_Carrier81_Faults_1" bit 2
   5204: 'Carrier 81 Drive: Error internal communications', class No Acknowledgement, trigger "DB302_HMI_Faults_Carrier81_Faults_1" bit 3
   5205: 'Carrier 81 Drive: Motor overtemperature', class No Acknowledgement, trigger "DB302_HMI_Faults_Carrier81_Faults_1" bit 4
   5206: 'Carrier 81 Drive: Motor overcurrent', class No Acknowledgement, trigger "DB302_HMI_Faults_Carrier81_Faults_1" bit 5
   5207: 'Carrier 81 Drive: Infeed or power unit not ready', class No Acknowledgement, trigger "DB302_HMI_Faults_Carrier81_Faults_1" bit 6
   5208: 'Carrier 81 Drive: Short-circuit/ground fault detected', class No Acknowledgement, trigger "DB302_HMI_Faults_Carrier81_Faults_1" bit 7
   5209: 'Carrier 81 Drive: PROFINET Setpoint timeout', class No Acknowledgement, trigger "DB302_HMI_Faults_Carrier81_Faults_1" bit 8
   5210: 'Carrier 81 Power unit: Overcurrent', class No Acknowledgement, trigger "DB302_HMI_Faults_Carrier81_Faults_1" bit 9
   5211: 'Carrier 81 Power unit: DC link voltage overvoltage', class No Acknowledgement, trigger "DB302_HMI_Faults_Carrier81_Faults_1" bit 10
   5212: 'Carrier 81 Power unit: DC link voltage undervoltage', class No Acknowledgement, trigger "DB302_HMI_Faults_Carrier81_Faults_1" bit 11
   5213: 'Carrier 81 Power unit: Line phase failure in main circuit', class No Acknowledgement, trigger "DB302_HMI_Faults_Carrier81_Faults_1" bit 12
   5214: 'Carrier 81 Power unit: Phase failure motor cable', class No Acknowledgement, trigger "DB302_HMI_Faults_Carrier81_Faults_1" bit 13
   5215: 'Carrier 81 Power unit: Ground fault', class No Acknowledgement, trigger "DB302_HMI_Faults_Carrier81_Faults_1" bit 14
   5216: 'Spare_Fault_5216', class No Acknowledgement, trigger "DB302_HMI_Faults_Carrier81_Faults_1" bit 15
   5217: 'Carrier 81 Motion Off Fault', class No Acknowledgement, trigger "DB302_HMI_Faults_Carrier81_Faults_2" bit 0
   5218: 'Carrier 81 Motion On Fault', class No Acknowledgement, trigger "DB302_HMI_Faults_Carrier81_Faults_2" bit 1
   5219: 'Carrier 81 Spacing Fault', class No Acknowledgement, trigger "DB302_HMI_Faults_Carrier81_Faults_2" bit 2
   5220: 'Carrier 81 Duplicate Carrier Number Fault', class No Acknowledgement, trigger "DB302_HMI_Faults_Carrier81_Faults_2" bit 3
   5221: 'Spare_Fault_5221', class No Acknowledgement, trigger "DB302_HMI_Faults_Carrier81_Faults_2" bit 4
   5222: 'Spare_Fault_5222', class No Acknowledgement, trigger "DB302_HMI_Faults_Carrier81_Faults_2" bit 5
   5223: 'Spare_Fault_5223', class No Acknowledgement, trigger "DB302_HMI_Faults_Carrier81_Faults_2" bit 6
   5224: 'Spare_Fault_5224', class No Acknowledgement, trigger "DB302_HMI_Faults_Carrier81_Faults_2" bit 7
   5225: 'Spare_Fault_5225', class No Acknowledgement, trigger "DB302_HMI_Faults_Carrier81_Faults_2" bit 8
   5226: 'Spare_Fault_5226', class No Acknowledgement, trigger "DB302_HMI_Faults_Carrier81_Faults_2" bit 9
   5227: 'Spare_Fault_5227', class No Acknowledgement, trigger "DB302_HMI_Faults_Carrier81_Faults_2" bit 10
   5228: 'Spare_Fault_5228', class No Acknowledgement, trigger "DB302_HMI_Faults_Carrier81_Faults_2" bit 11
   5229: 'Spare_Fault_5229', class No Acknowledgement, trigger "DB302_HMI_Faults_Carrier81_Faults_2" bit 12
   5230: 'Spare_Fault_5230', class No Acknowledgement, trigger "DB302_HMI_Faults_Carrier81_Faults_2" bit 13
   5231: 'Spare_Fault_5231', class No Acknowledgement, trigger "DB302_HMI_Faults_Carrier81_Faults_2" bit 14
   5232: 'Spare_Fault_5232', class No Acknowledgement, trigger "DB302_HMI_Faults_Carrier81_Faults_2" bit 15
   5233: 'Spare_Fault_5233', class No Acknowledgement, trigger "DB302_HMI_Faults_Carrier81_Faults_3" bit 0
   5234: 'Spare_Fault_5234', class No Acknowledgement, trigger "DB302_HMI_Faults_Carrier81_Faults_3" bit 1
   5235: 'Spare_Fault_5235', class No Acknowledgement, trigger "DB302_HMI_Faults_Carrier81_Faults_3" bit 2
   5236: 'Spare_Fault_5236', class No Acknowledgement, trigger "DB302_HMI_Faults_Carrier81_Faults_3" bit 3
   5237: 'Spare_Fault_5237', class No Acknowledgement, trigger "DB302_HMI_Faults_Carrier81_Faults_3" bit 4
   5238: 'Spare_Fault_5238', class No Acknowledgement, trigger "DB302_HMI_Faults_Carrier81_Faults_3" bit 5
   5239: 'Spare_Fault_5239', class No Acknowledgement, trigger "DB302_HMI_Faults_Carrier81_Faults_3" bit 6
   5240: 'Spare_Fault_5240', class No Acknowledgement, trigger "DB302_HMI_Faults_Carrier81_Faults_3" bit 7
   5241: 'Spare_Fault_5241', class No Acknowledgement, trigger "DB302_HMI_Faults_Carrier81_Faults_3" bit 8
   5242: 'Spare_Fault_5242', class No Acknowledgement, trigger "DB302_HMI_Faults_Carrier81_Faults_3" bit 9
   5243: 'Spare_Fault_5243', class No Acknowledgement, trigger "DB302_HMI_Faults_Carrier81_Faults_3" bit 10
   5244: 'Spare_Fault_5244', class No Acknowledgement, trigger "DB302_HMI_Faults_Carrier81_Faults_3" bit 11
   5245: 'Spare_Fault_5245', class No Acknowledgement, trigger "DB302_HMI_Faults_Carrier81_Faults_3" bit 12
   5246: 'Spare_Fault_5246', class No Acknowledgement, trigger "DB302_HMI_Faults_Carrier81_Faults_3" bit 13
   5247: 'Spare_Fault_5247', class No Acknowledgement, trigger "DB302_HMI_Faults_Carrier81_Faults_3" bit 14
   5248: 'Spare_Fault_5248', class No Acknowledgement, trigger "DB302_HMI_Faults_Carrier81_Faults_3" bit 15
   5249: 'Carrier 82 Disconnect Open Power Fault DI11.0', class No Acknowledgement, trigger "DB302_HMI_Faults_Carrier82_Faults_0" bit 0
   5250: 'Carrier 82 Drive Profinet Comm Fault', class No Acknowledgement, trigger "DB302_HMI_Faults_Carrier82_Faults_0" bit 1
   5251: 'Carrier 82 Production Stop Not Reset', class No Acknowledgement, trigger "DB302_HMI_Faults_Carrier82_Faults_0" bit 2
   5252: 'Carrier 82 CB02122 Tripped', class No Acknowledgement, trigger "DB302_HMI_Faults_Carrier82_Faults_0" bit 3
   5253: 'Carrier 82 CB02123 Tripped', class No Acknowledgement, trigger "DB302_HMI_Faults_Carrier82_Faults_0" bit 4
   5254: 'Carrier 82 AUX1 CB Tripped', class No Acknowledgement, trigger "DB302_HMI_Faults_Carrier82_Faults_0" bit 5
   5255: 'Carrier 82 AUX2 CB Tripped', class No Acknowledgement, trigger "DB302_HMI_Faults_Carrier82_Faults_0" bit 6
   5256: 'Carrier 82 PLC Not Communicating', class No Acknowledgement, trigger "DB302_HMI_Faults_Carrier82_Faults_0" bit 7
   5257: 'Carrier 82 Safe Input Card Fault', class No Acknowledgement, trigger "DB302_HMI_Faults_Carrier82_Faults_0" bit 8
   5258: 'Carrier 82 Safe Output Card Fault', class No Acknowledgement, trigger "DB302_HMI_Faults_Carrier82_Faults_0" bit 9
   5259: 'Carrier 82 Standard Input Card Fault', class No Acknowledgement, trigger "DB302_HMI_Faults_Carrier82_Faults_0" bit 10
   5260: 'Carrier 82 Standard Output Card Fault', class No Acknowledgement, trigger "DB302_HMI_Faults_Carrier82_Faults_0" bit 11
   5261: 'Carrier 82 Encoder Position Fault', class No Acknowledgement, trigger "DB302_HMI_Faults_Carrier82_Faults_0" bit 12
   5262: 'Carrier 82 Encoder Internal Error', class No Acknowledgement, trigger "DB302_HMI_Faults_Carrier82_Faults_0" bit 13
   5263: 'Carrier 82 Encoder Comm Fault', class No Acknowledgement, trigger "DB302_HMI_Faults_Carrier82_Faults_0" bit 14
   5264: 'Carrier 82 HMI Comm Fault', class No Acknowledgement, trigger "DB302_HMI_Faults_Carrier82_Faults_0" bit 15
   5265: 'Carrier 82 Crash Detection Fault', class No Acknowledgement, trigger "DB302_HMI_Faults_Carrier82_Faults_1" bit 0
   5266: 'Carrier 82 Carrier Number Invalid', class No Acknowledgement, trigger "DB302_HMI_Faults_Carrier82_Faults_1" bit 1
   5267: 'Carrier 82 Drive: PROFINET configuration error', class No Acknowledgement, trigger "DB302_HMI_Faults_Carrier82_Faults_1" bit 2
   5268: 'Carrier 82 Drive: Error internal communications', class No Acknowledgement, trigger "DB302_HMI_Faults_Carrier82_Faults_1" bit 3
   5269: 'Carrier 82 Drive: Motor overtemperature', class No Acknowledgement, trigger "DB302_HMI_Faults_Carrier82_Faults_1" bit 4
   5270: 'Carrier 82 Drive: Motor overcurrent', class No Acknowledgement, trigger "DB302_HMI_Faults_Carrier82_Faults_1" bit 5
   5271: 'Carrier 82 Drive: Infeed or power unit not ready', class No Acknowledgement, trigger "DB302_HMI_Faults_Carrier82_Faults_1" bit 6
   5272: 'Carrier 82 Drive: Short-circuit/ground fault detected', class No Acknowledgement, trigger "DB302_HMI_Faults_Carrier82_Faults_1" bit 7
   5273: 'Carrier 82 Drive: PROFINET Setpoint timeout', class No Acknowledgement, trigger "DB302_HMI_Faults_Carrier82_Faults_1" bit 8
   5274: 'Carrier 82 Power unit: Overcurrent', class No Acknowledgement, trigger "DB302_HMI_Faults_Carrier82_Faults_1" bit 9
   5275: 'Carrier 82 Power unit: DC link voltage overvoltage', class No Acknowledgement, trigger "DB302_HMI_Faults_Carrier82_Faults_1" bit 10
   5276: 'Carrier 82 Power unit: DC link voltage undervoltage', class No Acknowledgement, trigger "DB302_HMI_Faults_Carrier82_Faults_1" bit 11
   5277: 'Carrier 82 Power unit: Line phase failure in main circuit', class No Acknowledgement, trigger "DB302_HMI_Faults_Carrier82_Faults_1" bit 12
   5278: 'Carrier 82 Power unit: Phase failure motor cable', class No Acknowledgement, trigger "DB302_HMI_Faults_Carrier82_Faults_1" bit 13
   5279: 'Carrier 82 Power unit: Ground fault', class No Acknowledgement, trigger "DB302_HMI_Faults_Carrier82_Faults_1" bit 14
   5280: 'Spare_Fault_5280', class No Acknowledgement, trigger "DB302_HMI_Faults_Carrier82_Faults_1" bit 15
   5281: 'Carrier 82 Motion Off Fault', class No Acknowledgement, trigger "DB302_HMI_Faults_Carrier82_Faults_2" bit 0
   5282: 'Carrier 82 Motion On Fault', class No Acknowledgement, trigger "DB302_HMI_Faults_Carrier82_Faults_2" bit 1
   5283: 'Carrier 82 Spacing Fault', class No Acknowledgement, trigger "DB302_HMI_Faults_Carrier82_Faults_2" bit 2
   5284: 'Carrier 82 Duplicate Carrier Number Fault', class No Acknowledgement, trigger "DB302_HMI_Faults_Carrier82_Faults_2" bit 3
   5285: 'Spare_Fault_5285', class No Acknowledgement, trigger "DB302_HMI_Faults_Carrier82_Faults_2" bit 4
   5286: 'Spare_Fault_5286', class No Acknowledgement, trigger "DB302_HMI_Faults_Carrier82_Faults_2" bit 5
   5287: 'Spare_Fault_5287', class No Acknowledgement, trigger "DB302_HMI_Faults_Carrier82_Faults_2" bit 6
   5288: 'Spare_Fault_5288', class No Acknowledgement, trigger "DB302_HMI_Faults_Carrier82_Faults_2" bit 7
   5289: 'Spare_Fault_5289', class No Acknowledgement, trigger "DB302_HMI_Faults_Carrier82_Faults_2" bit 8
   5290: 'Spare_Fault_5290', class No Acknowledgement, trigger "DB302_HMI_Faults_Carrier82_Faults_2" bit 9
   5291: 'Spare_Fault_5291', class No Acknowledgement, trigger "DB302_HMI_Faults_Carrier82_Faults_2" bit 10
   5292: 'Spare_Fault_5292', class No Acknowledgement, trigger "DB302_HMI_Faults_Carrier82_Faults_2" bit 11
   5293: 'Spare_Fault_5293', class No Acknowledgement, trigger "DB302_HMI_Faults_Carrier82_Faults_2" bit 12
   5294: 'Spare_Fault_5294', class No Acknowledgement, trigger "DB302_HMI_Faults_Carrier82_Faults_2" bit 13
   5295: 'Spare_Fault_5295', class No Acknowledgement, trigger "DB302_HMI_Faults_Carrier82_Faults_2" bit 14
   5296: 'Spare_Fault_5296', class No Acknowledgement, trigger "DB302_HMI_Faults_Carrier82_Faults_2" bit 15
   5297: 'Spare_Fault_5297', class No Acknowledgement, trigger "DB302_HMI_Faults_Carrier82_Faults_3" bit 0
   5298: 'Spare_Fault_5298', class No Acknowledgement, trigger "DB302_HMI_Faults_Carrier82_Faults_3" bit 1
   5299: 'Spare_Fault_5299', class No Acknowledgement, trigger "DB302_HMI_Faults_Carrier82_Faults_3" bit 2
   5300: 'Spare_Fault_5300', class No Acknowledgement, trigger "DB302_HMI_Faults_Carrier82_Faults_3" bit 3
   5301: 'Spare_Fault_5301', class No Acknowledgement, trigger "DB302_HMI_Faults_Carrier82_Faults_3" bit 4
   5302: 'Spare_Fault_5302', class No Acknowledgement, trigger "DB302_HMI_Faults_Carrier82_Faults_3" bit 5
   5303: 'Spare_Fault_5303', class No Acknowledgement, trigger "DB302_HMI_Faults_Carrier82_Faults_3" bit 6
   5304: 'Spare_Fault_5304', class No Acknowledgement, trigger "DB302_HMI_Faults_Carrier82_Faults_3" bit 7
   5305: 'Spare_Fault_5305', class No Acknowledgement, trigger "DB302_HMI_Faults_Carrier82_Faults_3" bit 8
   5306: 'Spare_Fault_5306', class No Acknowledgement, trigger "DB302_HMI_Faults_Carrier82_Faults_3" bit 9
   5307: 'Spare_Fault_5307', class No Acknowledgement, trigger "DB302_HMI_Faults_Carrier82_Faults_3" bit 10
   5308: 'Spare_Fault_5308', class No Acknowledgement, trigger "DB302_HMI_Faults_Carrier82_Faults_3" bit 11
   5309: 'Spare_Fault_5309', class No Acknowledgement, trigger "DB302_HMI_Faults_Carrier82_Faults_3" bit 12
   5310: 'Spare_Fault_5310', class No Acknowledgement, trigger "DB302_HMI_Faults_Carrier82_Faults_3" bit 13
   5311: 'Spare_Fault_5311', class No Acknowledgement, trigger "DB302_HMI_Faults_Carrier82_Faults_3" bit 14
   5312: 'Spare_Fault_5312', class No Acknowledgement, trigger "DB302_HMI_Faults_Carrier82_Faults_3" bit 15
   4: 'Wireless Access Point 3 Comm Fault', class No Acknowledgement, trigger "DB302_HMI_Faults_SDC_Faults_0" bit 3